REGION Network 37: Validation position reached with module correction
   RUNG wire#powerrail
      Contact( #TMP_xAlwaysON )
      wire#w1
      Contact( #STC_tPZD_Pos.tR.tZSW1.x10 )
      wire#w2
      P_Trig( #STC_tOS_PN.x7 )
      Contact( #STC_tEXT_DATA.tW.xModuleCorrect )
      Contact( #IN_xPositioning )
      { S7_Templates := "SrcType := DInt" } LT_Contact(in1 := #STC_tPROP.d4, in2 := DINT#0)
      S_Coil( #STC_tST.x7 )
   END_RUNG
   RUNG wire#w2
      Contact( #STC_tST.x11 )
      Contact( #STC_tEXT_DATA.tW.xModuleCorrect )
      Contact( #IN_xPositioning )
      { S7_Templates := "SrcType := DInt" } EQ_Contact(in1 := #STC_tPROP.d4, in2 := DINT#0)
      S_Coil( #STC_tST.x7 )
   END_RUNG
   RUNG wire#w1
      I_Contact( #STC_tUSER_DATA.tR.xReadyToMove )
      wire#w3
      R_Coil( #STC_tST.x7 )
   END_RUNG
   RUNG wire#w1
      I_Contact( #IN_xPositioning )
   END_RUNG wire#w3
   RUNG wire#w1
      I_Contact( #STC_tEXT_DATA.tW.xModuleCorrect )
   END_RUNG wire#w3
   RUNG wire#w1
      { S7_Templates := "SrcType := DInt" } GT_Contact(in1 := #STC_tPROP.d4, in2 := DINT#0)
   END_RUNG wire#w3
   // the same network as SCL:
   #_w1 := #TMP_xAlwaysON AND #STC_tPZD_Pos.tR.tZSW1.x10;
   #_w2 := #_w1 AND NOT #STC_tOS_PN.x7;   // rising edge
   #STC_tOS_PN.x7 := #_w1;
   IF #_w2 AND #STC_tEXT_DATA.tW.xModuleCorrect AND #IN_xPositioning AND (#STC_tPROP.d4 < DINT#0) THEN
       #STC_tST.x7 := TRUE;
   END_IF;
   IF #_w1 AND #STC_tST.x11 AND #STC_tEXT_DATA.tW.xModuleCorrect AND #IN_xPositioning AND (#STC_tPROP.d4 = DINT#0) THEN
       #STC_tST.x7 := TRUE;
   END_IF;
   IF #TMP_xAlwaysON AND (NOT #STC_tUSER_DATA.tR.xReadyToMove OR NOT #IN_xPositioning OR NOT #STC_tEXT_DATA.tW.xModuleCorrect OR (#STC_tPROP.d4 > DINT#0)) THEN
       #STC_tST.x7 := FALSE;
   END_IF;
END_REGION

REGION Network 38: Positioning reached
   RUNG wire#powerrail
      Contact( #STC_tUSER_DATA.tR.xReadyToMove )
      Contact( #IN_xPositioning )
      Contact( #STC_tPZD_Pos.tR.tZSW1.x10 )
      wire#w1
      { S7_Templates := "SrcType := DInt" } GE_Contact(in1 := #STC_tPROP.d4, in2 := #TMP_dActualPosMin_cmm)
      { S7_Templates := "SrcType := DInt" } LE_Contact(in1 := #STC_tPROP.d4, in2 := #TMP_dActualPosMax_cmm)
      wire#w2
      Contact( #STC_tPZD_Pos.tR.tPOS_ZSW2.x2 )
      I_Contact( #STC_tPZD_Pos.tR.tPOS_ZSW2.x15 )
      I_Contact( #STC_tPZD_Pos.tW.tSTW1.x6 )
      I_Contact( #STC_tPZD_Pos.tR.tZSW1.x12 )
      Coil( #TMP_x )
   END_RUNG
   RUNG wire#w1
      Contact( #STC_tUSER_DATA.tW.xRelativePosition )
   END_RUNG wire#w2
   RUNG wire#w1
      { S7_Templates := "SrcType := DInt" } LT_Contact(in1 := #STC_tPROP.d4, in2 := 0)
   END_RUNG wire#w2
   RUNG wire#w1
      Contact( #STC_tST.x7 )
   END_RUNG wire#w2
   // the same network as SCL:
   #TMP_x := #STC_tUSER_DATA.tR.xReadyToMove AND #IN_xPositioning AND #STC_tPZD_Pos.tR.tZSW1.x10 AND (((#STC_tPROP.d4 >= #TMP_dActualPosMin_cmm) AND (#STC_tPROP.d4 <= #TMP_dActualPosMax_cmm)) OR #STC_tUSER_DATA.tW.xRelativePosition OR (#STC_tPROP.d4 < 0) OR #STC_tST.x7) AND #STC_tPZD_Pos.tR.tPOS_ZSW2.x2 AND NOT #STC_tPZD_Pos.tR.tPOS_ZSW2.x15 AND NOT #STC_tPZD_Pos.tW.tSTW1.x6 AND NOT #STC_tPZD_Pos.tR.tZSW1.x12;
END_REGION

REGION Network 39: Positioning reached
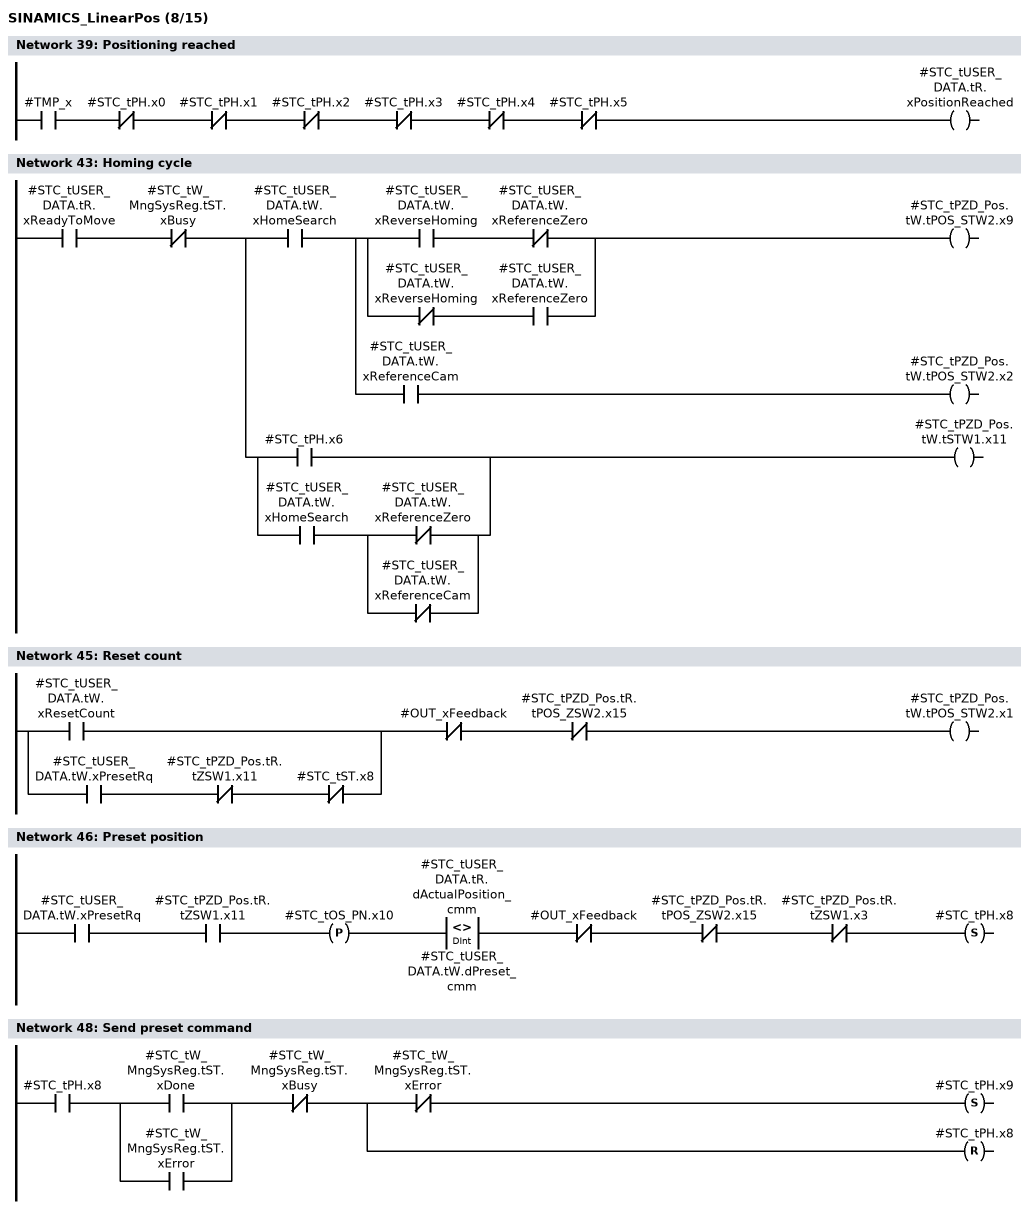
   RUNG wire#powerrail
      Contact( #TMP_x )
      I_Contact( #STC_tPH.x0 )
      I_Contact( #STC_tPH.x1 )
      I_Contact( #STC_tPH.x2 )
      I_Contact( #STC_tPH.x3 )
      I_Contact( #STC_tPH.x4 )
      I_Contact( #STC_tPH.x5 )
      Coil( #STC_tUSER_DATA.tR.xPositionReached )
   END_RUNG
   // the same network as SCL:
   #STC_tUSER_DATA.tR.xPositionReached := #TMP_x AND NOT #STC_tPH.x0 AND NOT #STC_tPH.x1 AND NOT #STC_tPH.x2 AND NOT #STC_tPH.x3 AND NOT #STC_tPH.x4 AND NOT #STC_tPH.x5;
END_REGION

REGION Network 40: #####_HOMING_CYCLE_#####
END_REGION

REGION Network 41 (STL): Send homing preset
         A     #STC_tUSER_DATA.tW.xHomeSearch;
         AN    #STC_tPZD_Pos.tW.tSTW1.x11;
         JCN   PrH0;
         =     #STC_tW_MngSysReg.tST.xWrite_Request;

         L     #STC_tSYS_DATA.iPosPZD_MM;
         SLW   8;
         L     W#16#2;
         OW;
         T     #STC_tW_MngSysReg.tDATA.wRequest_refere_RequestID;
         L     #STC_tSYS_DATA.iPosPZD_MM;
         SLW   8;
         L     W#16#1;
         OW;
         T     #STC_tW_MngSysReg.tDATA.wAxis_NoOfParameters;
         L     W#16#1001;
         T     #STC_tW_MngSysReg.tDATA.wAttribute_NoOfElements;
         L     2599;
         T     #STC_tW_MngSysReg.tDATA.iParameter_number;
         L     W#16#0;
         T     #STC_tW_MngSysReg.tDATA.wSubindex;
         L     W#16#4301;
         T     #STC_tW_MngSysReg.tDATA.wFormat_NoOfValue;
         L     #STC_tSYS_DATA.iDiagAddress;
         T     #STC_tW_MngSysReg.tST.ID;
         L     47;
         T     #STC_tW_MngSysReg.tST.dINDEX;
         L     16;
         T     #STC_tW_MngSysReg.tST.uiLEN;

         L     #STC_tUSER_DATA.tW.dPreset_cmm;
   //      L     DINT#10
   //      *D
         T     #STC_tW_MngSysReg.tDATA.dwRegisterValue;

         CALL  #STC_tWriteRecord
         ( REQ    := #STC_tW_MngSysReg.tST.xWrite_Request,
           ID     := #STC_tW_MngSysReg.tST.ID,
           INDEX  := #STC_tW_MngSysReg.tST.dINDEX,
           LEN    := #STC_tW_MngSysReg.tST.uiLEN,
           DONE   := #STC_tW_MngSysReg.tST.xDone,
           BUSY   := #STC_tW_MngSysReg.tST.xBusy,
           ERROR  := #STC_tW_MngSysReg.tST.xError,
           STATUS := #STC_tW_MngSysReg.tST.dwSTATUS,
           RECORD := #STC_tW_MngSysReg.tDATA
         );
   PrH0: NOP   0;
END_REGION

REGION Network 42 (STL): Error during Send homing preset
         A     #STC_tW_MngSysReg.tST.xError;
         L     34;
         JC    Err;
END_REGION

REGION Network 43: Homing cycle
   RUNG wire#powerrail
      Contact( #STC_tUSER_DATA.tR.xReadyToMove )
      I_Contact( #STC_tW_MngSysReg.tST.xBusy )
      wire#w1
      Contact( #STC_tUSER_DATA.tW.xHomeSearch )
      wire#w2
      Contact( #STC_tUSER_DATA.tW.xReverseHoming )
      I_Contact( #STC_tUSER_DATA.tW.xReferenceZero )
      wire#w3
      Coil( #STC_tPZD_Pos.tW.tPOS_STW2.x9 )
   END_RUNG
   RUNG wire#w2
      I_Contact( #STC_tUSER_DATA.tW.xReverseHoming )
      Contact( #STC_tUSER_DATA.tW.xReferenceZero )
   END_RUNG wire#w3
   RUNG wire#w2
      Contact( #STC_tUSER_DATA.tW.xReferenceCam )
      Coil( #STC_tPZD_Pos.tW.tPOS_STW2.x2 )
   END_RUNG
   RUNG wire#w1
      Contact( #STC_tPH.x6 )
      wire#w4
      Coil( #STC_tPZD_Pos.tW.tSTW1.x11 )
   END_RUNG
   RUNG wire#w1
      Contact( #STC_tUSER_DATA.tW.xHomeSearch )
      wire#w5
      I_Contact( #STC_tUSER_DATA.tW.xReferenceZero )
   END_RUNG wire#w4
   RUNG wire#w5
      I_Contact( #STC_tUSER_DATA.tW.xReferenceCam )
   END_RUNG wire#w4
   // the same network as SCL:
   #_w1 := #STC_tUSER_DATA.tR.xReadyToMove AND NOT #STC_tW_MngSysReg.tST.xBusy;
   #_w2 := #_w1 AND #STC_tUSER_DATA.tW.xHomeSearch;
   #STC_tPZD_Pos.tW.tPOS_STW2.x9 := #_w2 AND ((#STC_tUSER_DATA.tW.xReverseHoming AND NOT #STC_tUSER_DATA.tW.xReferenceZero) OR (NOT #STC_tUSER_DATA.tW.xReverseHoming AND #STC_tUSER_DATA.tW.xReferenceZero));
   #STC_tPZD_Pos.tW.tPOS_STW2.x2 := #_w2 AND #STC_tUSER_DATA.tW.xReferenceCam;
   #STC_tPZD_Pos.tW.tSTW1.x11 := #_w1 AND (#STC_tPH.x6 OR (#STC_tUSER_DATA.tW.xHomeSearch AND (NOT #STC_tUSER_DATA.tW.xReferenceZero OR NOT #STC_tUSER_DATA.tW.xReferenceCam)));
END_REGION

REGION Network 44: #####_PRESET_ACTUAL_POSITION_#####
END_REGION

REGION Network 45: Reset count
   RUNG wire#powerrail
      Contact( #STC_tUSER_DATA.tW.xResetCount )
      wire#w1
      I_Contact( #OUT_xFeedback )
      I_Contact( #STC_tPZD_Pos.tR.tPOS_ZSW2.x15 )
      Coil( #STC_tPZD_Pos.tW.tPOS_STW2.x1 )
   END_RUNG
   RUNG wire#powerrail
      Contact( #STC_tUSER_DATA.tW.xPresetRq )
      I_Contact( #STC_tPZD_Pos.tR.tZSW1.x11 )
      I_Contact( #STC_tST.x8 )
   END_RUNG wire#w1
   // the same network as SCL:
   #STC_tPZD_Pos.tW.tPOS_STW2.x1 := (#STC_tUSER_DATA.tW.xResetCount OR (#STC_tUSER_DATA.tW.xPresetRq AND NOT #STC_tPZD_Pos.tR.tZSW1.x11 AND NOT #STC_tST.x8)) AND NOT #OUT_xFeedback AND NOT #STC_tPZD_Pos.tR.tPOS_ZSW2.x15;
END_REGION

REGION Network 46: Preset position
   RUNG wire#powerrail
      Contact( #STC_tUSER_DATA.tW.xPresetRq )
      Contact( #STC_tPZD_Pos.tR.tZSW1.x11 )
      P_Trig( #STC_tOS_PN.x10 )
      { S7_Templates := "SrcType := DInt" } NE_Contact(in1 := #STC_tUSER_DATA.tR.dActualPosition_cmm, in2 := #STC_tUSER_DATA.tW.dPreset_cmm)
      I_Contact( #OUT_xFeedback )
      I_Contact( #STC_tPZD_Pos.tR.tPOS_ZSW2.x15 )
      I_Contact( #STC_tPZD_Pos.tR.tZSW1.x3 )
      S_Coil( #STC_tPH.x8 )
   END_RUNG
   // the same network as SCL:
   #_w1 := #STC_tUSER_DATA.tW.xPresetRq AND #STC_tPZD_Pos.tR.tZSW1.x11;
   #_w2 := #_w1 AND NOT #STC_tOS_PN.x10;   // rising edge
   #STC_tOS_PN.x10 := #_w1;
   IF #_w2 AND (#STC_tUSER_DATA.tR.dActualPosition_cmm <> #STC_tUSER_DATA.tW.dPreset_cmm) AND NOT #OUT_xFeedback AND NOT #STC_tPZD_Pos.tR.tPOS_ZSW2.x15 AND NOT #STC_tPZD_Pos.tR.tZSW1.x3 THEN
       #STC_tPH.x8 := TRUE;
   END_IF;
END_REGION

REGION Network 47 (STL): Send encoder value
         A     #STC_tPH.x8;
         JCN   PrE0;
         =     #STC_tW_MngSysReg.tST.xWrite_Request;

         L     #STC_tSYS_DATA.iPosPZD_MM;
         +     10;
         SLW   8;
         L     W#16#2;
         OW;
         T     #STC_tW_MngSysReg.tDATA.wRequest_refere_RequestID;
         L     #STC_tSYS_DATA.iPosPZD_MM;
         SLW   8;
         L     W#16#1;
         OW;
         T     #STC_tW_MngSysReg.tDATA.wAxis_NoOfParameters;
         L     W#16#1001;
         T     #STC_tW_MngSysReg.tDATA.wAttribute_NoOfElements;
         L     2599;
         T     #STC_tW_MngSysReg.tDATA.iParameter_number;
         L     W#16#0;
         T     #STC_tW_MngSysReg.tDATA.wSubindex;
         L     W#16#4301;
         T     #STC_tW_MngSysReg.tDATA.wFormat_NoOfValue;
         L     #STC_tSYS_DATA.iDiagAddress;
         T     #STC_tW_MngSysReg.tST.ID;
         L     47;
         T     #STC_tW_MngSysReg.tST.dINDEX;
         L     16;
         T     #STC_tW_MngSysReg.tST.uiLEN;

         L     #STC_tUSER_DATA.tW.dPreset_cmm;
   //  L     DINT#10
   //  *D
         T     #STC_tW_MngSysReg.tDATA.dwRegisterValue;

         CALL  #STC_tWriteRecord
         ( REQ    := #STC_tW_MngSysReg.tST.xWrite_Request,
           ID     := #STC_tW_MngSysReg.tST.ID,
           INDEX  := #STC_tW_MngSysReg.tST.dINDEX,
           LEN    := #STC_tW_MngSysReg.tST.uiLEN,
           DONE   := #STC_tW_MngSysReg.tST.xDone,
           BUSY   := #STC_tW_MngSysReg.tST.xBusy,
           ERROR  := #STC_tW_MngSysReg.tST.xError,
           STATUS := #STC_tW_MngSysReg.tST.dwSTATUS,
           RECORD := #STC_tW_MngSysReg.tDATA
         );
   PrE0: NOP   0;
END_REGION

REGION Network 48: Send preset command
   RUNG wire#powerrail
      Contact( #STC_tPH.x8 )
      wire#w1
      Contact( #STC_tW_MngSysReg.tST.xDone )
      wire#w2
      I_Contact( #STC_tW_MngSysReg.tST.xBusy )
      wire#w3
      I_Contact( #STC_tW_MngSysReg.tST.xError )
      S_Coil( #STC_tPH.x9 )
   END_RUNG
   RUNG wire#w1
      Contact( #STC_tW_MngSysReg.tST.xError )
   END_RUNG wire#w2
   RUNG wire#w3
      R_Coil( #STC_tPH.x8 )
   END_RUNG
   // the same network as SCL:
   #_w1 := #STC_tPH.x8 AND (#STC_tW_MngSysReg.tST.xDone OR #STC_tW_MngSysReg.tST.xError) AND NOT #STC_tW_MngSysReg.tST.xBusy;
   IF #_w1 AND NOT #STC_tW_MngSysReg.tST.xError THEN #STC_tPH.x9 := TRUE; END_IF;
   IF #_w1 THEN #STC_tPH.x8 := FALSE; END_IF;
END_REGION

REGION Network 49 (STL): Error during send ecoder value
         A     #STC_tW_MngSysReg.tST.xError;
         L     30;
         JC    Err;
END_REGION

REGION Network 50 (STL): Send preset command
         A     #STC_tPH.x9;
         JCN   PrE1;
         =     #STC_tW_MngSysReg.tST.xWrite_Request;

         L     #STC_tSYS_DATA.iPosPZD_MM;
         +     20;
         SLW   8;
         L     W#16#2;
         OW;
         T     #STC_tW_MngSysReg.tDATA.wRequest_refere_RequestID;
         L     #STC_tSYS_DATA.iPosPZD_MM;
         SLW   8;
         L     W#16#1;
         OW;
         T     #STC_tW_MngSysReg.tDATA.wAxis_NoOfParameters;
         L     W#16#1001;
         T     #STC_tW_MngSysReg.tDATA.wAttribute_NoOfElements;
         L     2507;
         T     #STC_tW_MngSysReg.tDATA.iParameter_number;
         L     #STC_tSYS_DATA.iEncNumb;
         T     #STC_tW_MngSysReg.tDATA.wSubindex;
         L     W#16#4201;
         T     #STC_tW_MngSysReg.tDATA.wFormat_NoOfValue;
         L     #STC_tSYS_DATA.iDiagAddress;
         T     #STC_tW_MngSysReg.tST.ID;
         L     47;
         T     #STC_tW_MngSysReg.tST.dINDEX;
         L     14;
         T     #STC_tW_MngSysReg.tST.uiLEN;

         L     DINT#2;
         SLD   16;
         T     #STC_tW_MngSysReg.tDATA.dwRegisterValue;

         CALL  #STC_tWriteRecord
         ( REQ    := #STC_tW_MngSysReg.tST.xWrite_Request,
           ID     := #STC_tW_MngSysReg.tST.ID,
           INDEX  := #STC_tW_MngSysReg.tST.dINDEX,
           LEN    := #STC_tW_MngSysReg.tST.uiLEN,
           DONE   := #STC_tW_MngSysReg.tST.xDone,
           BUSY   := #STC_tW_MngSysReg.tST.xBusy,
           ERROR  := #STC_tW_MngSysReg.tST.xError,
           STATUS := #STC_tW_MngSysReg.tST.dwSTATUS,
           RECORD := #STC_tW_MngSysReg.tDATA
         );
   PrE1: NOP   0;
END_REGION

REGION Network 51: Send saving preset command
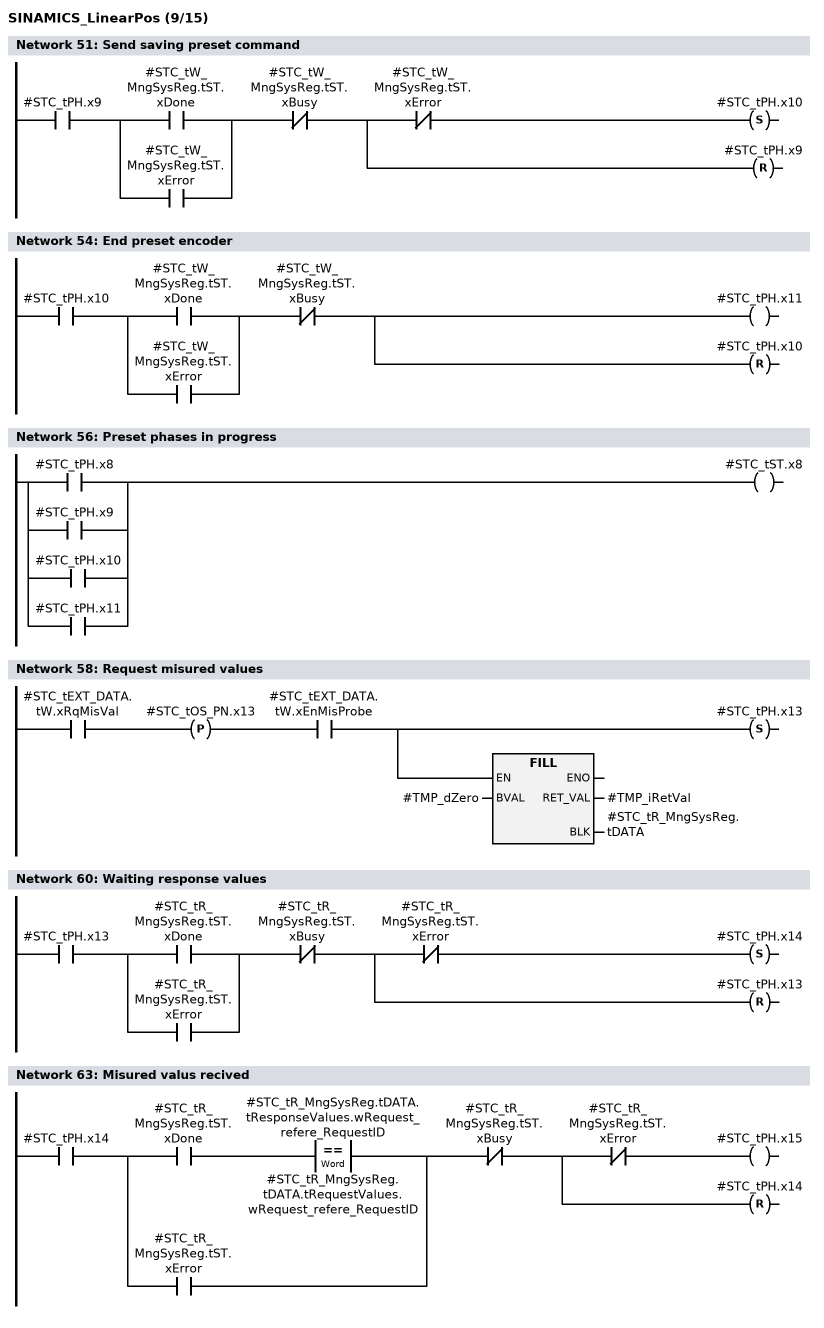
   RUNG wire#powerrail
      Contact( #STC_tPH.x9 )
      wire#w1
      Contact( #STC_tW_MngSysReg.tST.xDone )
      wire#w2
      I_Contact( #STC_tW_MngSysReg.tST.xBusy )
      wire#w3
      I_Contact( #STC_tW_MngSysReg.tST.xError )
      S_Coil( #STC_tPH.x10 )
   END_RUNG
   RUNG wire#w1
      Contact( #STC_tW_MngSysReg.tST.xError )
   END_RUNG wire#w2
   RUNG wire#w3
      R_Coil( #STC_tPH.x9 )
   END_RUNG
   // the same network as SCL:
   #_w1 := #STC_tPH.x9 AND (#STC_tW_MngSysReg.tST.xDone OR #STC_tW_MngSysReg.tST.xError) AND NOT #STC_tW_MngSysReg.tST.xBusy;
   IF #_w1 AND NOT #STC_tW_MngSysReg.tST.xError THEN #STC_tPH.x10 := TRUE; END_IF;
   IF #_w1 THEN #STC_tPH.x9 := FALSE; END_IF;
END_REGION

REGION Network 52 (STL): Error during preset command
         A     #STC_tW_MngSysReg.tST.xError;
         L     31;
         JC    Err;
END_REGION

REGION Network 53 (STL): Send saving preset command
         A     #STC_tPH.x10;
         JCN   PrE2;
         =     #STC_tW_MngSysReg.tST.xWrite_Request;

         L     #STC_tSYS_DATA.iPosPZD_MM;
         +     30;
         SLW   8;
         L     W#16#2;
         OW;
         T     #STC_tW_MngSysReg.tDATA.wRequest_refere_RequestID;
         L     #STC_tSYS_DATA.iPosPZD_CU;
         SLW   8;
         L     W#16#1;
         OW;
         T     #STC_tW_MngSysReg.tDATA.wAxis_NoOfParameters;
         L     W#16#1001;
         T     #STC_tW_MngSysReg.tDATA.wAttribute_NoOfElements;
         L     977;
         T     #STC_tW_MngSysReg.tDATA.iParameter_number;
         L     W#16#0;
         T     #STC_tW_MngSysReg.tDATA.wSubindex;
         L     W#16#4201;
         T     #STC_tW_MngSysReg.tDATA.wFormat_NoOfValue;
         L     #STC_tSYS_DATA.iDiagAddress;
         T     #STC_tW_MngSysReg.tST.ID;
         L     47;
         T     #STC_tW_MngSysReg.tST.dINDEX;
         L     14;
         T     #STC_tW_MngSysReg.tST.uiLEN;

         L     DINT#1;
         SLD   16;
         T     #STC_tW_MngSysReg.tDATA.dwRegisterValue;

         CALL  #STC_tWriteRecord
         ( REQ    := #STC_tW_MngSysReg.tST.xWrite_Request,
           ID     := #STC_tW_MngSysReg.tST.ID,
           INDEX  := #STC_tW_MngSysReg.tST.dINDEX,
           LEN    := #STC_tW_MngSysReg.tST.uiLEN,
           DONE   := #STC_tW_MngSysReg.tST.xDone,
           BUSY   := #STC_tW_MngSysReg.tST.xBusy,
           ERROR  := #STC_tW_MngSysReg.tST.xError,
           STATUS := #STC_tW_MngSysReg.tST.dwSTATUS,
           RECORD := #STC_tW_MngSysReg.tDATA
         );
   PrE2: NOP   0;
END_REGION

REGION Network 54: End preset encoder
   RUNG wire#powerrail
      Contact( #STC_tPH.x10 )
      wire#w1
      Contact( #STC_tW_MngSysReg.tST.xDone )
      wire#w2
      I_Contact( #STC_tW_MngSysReg.tST.xBusy )
      wire#w3
      Coil( #STC_tPH.x11 )
   END_RUNG
   RUNG wire#w1
      Contact( #STC_tW_MngSysReg.tST.xError )
   END_RUNG wire#w2
   RUNG wire#w3
      R_Coil( #STC_tPH.x10 )
   END_RUNG
   // the same network as SCL:
   #STC_tPH.x11 := #STC_tPH.x10 AND (#STC_tW_MngSysReg.tST.xDone OR #STC_tW_MngSysReg.tST.xError) AND NOT #STC_tW_MngSysReg.tST.xBusy;
   IF #STC_tPH.x11 THEN #STC_tPH.x10 := FALSE; END_IF;
END_REGION

REGION Network 55 (STL): Error during saving preset command
         A     #STC_tW_MngSysReg.tST.xError;
         L     32;
         JC    Err;
END_REGION

REGION Network 56: Preset phases in progress
   RUNG wire#powerrail
      Contact( #STC_tPH.x8 )
      wire#w1
      Coil( #STC_tST.x8 )
   END_RUNG
   RUNG wire#powerrail
      Contact( #STC_tPH.x9 )
   END_RUNG wire#w1
   RUNG wire#powerrail
      Contact( #STC_tPH.x10 )
   END_RUNG wire#w1
   RUNG wire#powerrail
      Contact( #STC_tPH.x11 )
   END_RUNG wire#w1
   // the same network as SCL:
   #STC_tST.x8 := #STC_tPH.x8 OR #STC_tPH.x9 OR #STC_tPH.x10 OR #STC_tPH.x11;
END_REGION

REGION Network 57: #####_READING_MISURED_VALUES_#####
END_REGION

REGION Network 58: Request misured values
   #_w1 := #STC_tEXT_DATA.tW.xRqMisVal AND NOT #STC_tOS_PN.x13;   // rising edge
   #STC_tOS_PN.x13 := #STC_tEXT_DATA.tW.xRqMisVal;
   IF #_w1 AND #STC_tEXT_DATA.tW.xEnMisProbe THEN
       #STC_tPH.x13 := TRUE;
       #TMP_iRetVal := FILL(BVAL := #TMP_dZero, BLK => #STC_tR_MngSysReg.tDATA);
   END_IF;
END_REGION

REGION Network 59 (STL): Send request misured values
         A     #STC_tPH.x13;
         JCN   RdV1;
         =     #STC_tR_MngSysReg.tST.xRead_Request;

         L     #STC_tSYS_DATA.iPosPZD_MM;
         +     40;
         SLW   8;
         L     W#16#1;
         OW;
         T     #STC_tR_MngSysReg.tDATA.tRequestValues.wRequest_refere_RequestID;
         L     #STC_tSYS_DATA.iPosPZD_MM;
         SLW   8;
         L     W#16#C;
         OW;
         T     #STC_tR_MngSysReg.tDATA.tRequestValues.wAxis_NoOfParameters;
         L     W#16#1000;
         T     #STC_tR_MngSysReg.tDATA.tRequestValues.wAttribute_NoOfElements_1;
         L     21700;
         T     #STC_tR_MngSysReg.tDATA.tRequestValues.iParameter_number_1;
         L     W#16#0;
         T     #STC_tR_MngSysReg.tDATA.tRequestValues.wSubindex_1;

         L     W#16#1000;
         T     #STC_tR_MngSysReg.tDATA.tRequestValues.wAttribute_NoOfElements_2;
         L     21701;
         T     #STC_tR_MngSysReg.tDATA.tRequestValues.iParameter_number_2;
         L     W#16#0;
         T     #STC_tR_MngSysReg.tDATA.tRequestValues.wSubindex_2;

         L     W#16#1000;
         T     #STC_tR_MngSysReg.tDATA.tRequestValues.wAttribute_NoOfElements_3;
         L     21702;
         T     #STC_tR_MngSysReg.tDATA.tRequestValues.iParameter_number_3;
         L     W#16#0;
         T     #STC_tR_MngSysReg.tDATA.tRequestValues.wSubindex_3;

         L     W#16#1000;
         T     #STC_tR_MngSysReg.tDATA.tRequestValues.wAttribute_NoOfElements_4;
         L     21703;
         T     #STC_tR_MngSysReg.tDATA.tRequestValues.iParameter_number_4;
         L     W#16#0;
         T     #STC_tR_MngSysReg.tDATA.tRequestValues.wSubindex_4;

         L     W#16#1000;
         T     #STC_tR_MngSysReg.tDATA.tRequestValues.wAttribute_NoOfElements_5;
         L     21704;
         T     #STC_tR_MngSysReg.tDATA.tRequestValues.iParameter_number_5;
         L     W#16#0;
         T     #STC_tR_MngSysReg.tDATA.tRequestValues.wSubindex_5;

         L     W#16#1000;
         T     #STC_tR_MngSysReg.tDATA.tRequestValues.wAttribute_NoOfElements_6;
         L     21705;
         T     #STC_tR_MngSysReg.tDATA.tRequestValues.iParameter_number_6;
         L     W#16#0;
         T     #STC_tR_MngSysReg.tDATA.tRequestValues.wSubindex_6;

         L     W#16#1000;
         T     #STC_tR_MngSysReg.tDATA.tRequestValues.wAttribute_NoOfElements_7;
         L     21712;
         T     #STC_tR_MngSysReg.tDATA.tRequestValues.iParameter_number_7;
         L     W#16#0;
         T     #STC_tR_MngSysReg.tDATA.tRequestValues.wSubindex_7;

         L     W#16#1000;
         T     #STC_tR_MngSysReg.tDATA.tRequestValues.wAttribute_NoOfElements_8;
         L     21713;
         T     #STC_tR_MngSysReg.tDATA.tRequestValues.iParameter_number_8;
         L     W#16#0;
         T     #STC_tR_MngSysReg.tDATA.tRequestValues.wSubindex_8;

         L     W#16#1000;
         T     #STC_tR_MngSysReg.tDATA.tRequestValues.wAttribute_NoOfElements_9;
         L     21714;
         T     #STC_tR_MngSysReg.tDATA.tRequestValues.iParameter_number_9;
         L     W#16#0;
         T     #STC_tR_MngSysReg.tDATA.tRequestValues.wSubindex_9;

         L     W#16#1000;
         T     #STC_tR_MngSysReg.tDATA.tRequestValues.wAttribute_NoOfElement_10;
         L     21715;
         T     #STC_tR_MngSysReg.tDATA.tRequestValues.iParameter_number_10;
         L     W#16#0;
         T     #STC_tR_MngSysReg.tDATA.tRequestValues.wSubindex_10;

         L     W#16#1000;
         T     #STC_tR_MngSysReg.tDATA.tRequestValues.wAttribute_NoOfElement_11;
         L     21716;
         T     #STC_tR_MngSysReg.tDATA.tRequestValues.iParameter_number_11;
         L     W#16#0;
         T     #STC_tR_MngSysReg.tDATA.tRequestValues.wSubindex_11;

         L     W#16#1000;
         T     #STC_tR_MngSysReg.tDATA.tRequestValues.wAttribute_NoOfElement_12;
         L     21717;
         T     #STC_tR_MngSysReg.tDATA.tRequestValues.iParameter_number_12;
         L     W#16#0;
         T     #STC_tR_MngSysReg.tDATA.tRequestValues.wSubindex_12;

         L     #STC_tSYS_DATA.iDiagAddress;
         T     #STC_tR_MngSysReg.tST.ID;
         L     47;
         T     #STC_tR_MngSysReg.tST.dINDEX;
         L     76;
         T     #STC_tR_MngSysReg.tST.uiLEN;

         CALL  #STC_tWriteRecord
         ( REQ    := #STC_tR_MngSysReg.tST.xRead_Request,
           ID     := #STC_tR_MngSysReg.tST.ID,
           INDEX  := #STC_tR_MngSysReg.tST.dINDEX,
           LEN    := #STC_tR_MngSysReg.tST.uiLEN,
           DONE   := #STC_tR_MngSysReg.tST.xDone,
           BUSY   := #STC_tR_MngSysReg.tST.xBusy,
           ERROR  := #STC_tR_MngSysReg.tST.xError,
           STATUS := #STC_tR_MngSysReg.tST.dwSTATUS,
           RECORD := #STC_tR_MngSysReg.tDATA.tRequestValues
         );

   RdV1: NOP   0;
END_REGION

REGION Network 60: Waiting response values
   RUNG wire#powerrail
      Contact( #STC_tPH.x13 )
      wire#w1
      Contact( #STC_tR_MngSysReg.tST.xDone )
      wire#w2
      I_Contact( #STC_tR_MngSysReg.tST.xBusy )
      wire#w3
      I_Contact( #STC_tR_MngSysReg.tST.xError )
      S_Coil( #STC_tPH.x14 )
   END_RUNG
   RUNG wire#w1
      Contact( #STC_tR_MngSysReg.tST.xError )
   END_RUNG wire#w2
   RUNG wire#w3
      R_Coil( #STC_tPH.x13 )
   END_RUNG
   // the same network as SCL:
   #_w1 := #STC_tPH.x13 AND (#STC_tR_MngSysReg.tST.xDone OR #STC_tR_MngSysReg.tST.xError) AND NOT #STC_tR_MngSysReg.tST.xBusy;
   IF #_w1 AND NOT #STC_tR_MngSysReg.tST.xError THEN #STC_tPH.x14 := TRUE; END_IF;
   IF #_w1 THEN #STC_tPH.x13 := FALSE; END_IF;
END_REGION

REGION Network 61 (STL): Error during waiting response values
         A     #STC_tR_MngSysReg.tST.xError;
         L     40;
         JC    Err;
END_REGION

REGION Network 62 (STL): Send response misured values
         A     #STC_tPH.x14;
         JCN   RdV2;
         AN    #STC_tR_MngSysReg.tST.xBusy;
         =     #STC_tR_MngSysReg.tST.xRead_Request;

         L     #STC_tSYS_DATA.iDiagAddress;
         T     #STC_tR_MngSysReg.tST.ID;
         L     47;
         T     #STC_tR_MngSysReg.tST.dINDEX;
         L     76;
         T     #STC_tR_MngSysReg.tST.uiMLEN;

         CALL  #STC_tReadRecord
         ( REQ    := #STC_tR_MngSysReg.tST.xRead_Request,
           ID     := #STC_tR_MngSysReg.tST.ID,
           INDEX  := #STC_tR_MngSysReg.tST.dINDEX,
           MLEN   := #STC_tR_MngSysReg.tST.uiMLEN,
           VALID  := #STC_tR_MngSysReg.tST.xDone,
           BUSY   := #STC_tR_MngSysReg.tST.xBusy,
           ERROR  := #STC_tR_MngSysReg.tST.xError,
           STATUS := #STC_tR_MngSysReg.tST.dwSTATUS,
           LEN    := #STC_tR_MngSysReg.tST.uiLEN,
           RECORD := #STC_tR_MngSysReg.tDATA.tResponseValues
         );

         L     #STC_tR_MngSysReg.tDATA.tResponseValues.wRequest_refere_RequestID;
         L     W#16#FF7F;
         AW;
         T     #STC_tR_MngSysReg.tDATA.tResponseValues.wRequest_refere_RequestID;

   RdV2: NOP   0;
END_REGION

REGION Network 63: Misured valus recived
   RUNG wire#powerrail
      Contact( #STC_tPH.x14 )
      wire#w1
      Contact( #STC_tR_MngSysReg.tST.xDone )
      { S7_Templates := "SrcType := Word" } EQ_Contact(in1 := #STC_tR_MngSysReg.tDATA.tResponseValues.wRequest_refere_RequestID, in2 := #STC_tR_MngSysReg.tDATA.tRequestValues.wRequest_refere_RequestID)
      wire#w2
      I_Contact( #STC_tR_MngSysReg.tST.xBusy )
      wire#w3
      I_Contact( #STC_tR_MngSysReg.tST.xError )
      Coil( #STC_tPH.x15 )
   END_RUNG
   RUNG wire#w1
      Contact( #STC_tR_MngSysReg.tST.xError )
   END_RUNG wire#w2
   RUNG wire#w3
      R_Coil( #STC_tPH.x14 )
   END_RUNG
   // the same network as SCL:
   #_w1 := #STC_tPH.x14 AND ((#STC_tR_MngSysReg.tST.xDone AND (#STC_tR_MngSysReg.tDATA.tResponseValues.wRequest_refere_RequestID = #STC_tR_MngSysReg.tDATA.tRequestValues.wRequest_refere_RequestID)) OR #STC_tR_MngSysReg.tST.xError) AND NOT #STC_tR_MngSysReg.tST.xBusy;
   #STC_tPH.x15 := #_w1 AND NOT #STC_tR_MngSysReg.tST.xError;
   IF #_w1 THEN #STC_tPH.x14 := FALSE; END_IF;
END_REGION

REGION Network 64 (STL): Error during misured valus recived
         A     #STC_tR_MngSysReg.tST.xError;
         L     41;
         JC    Err;
END_REGION

REGION Network 65: Save data
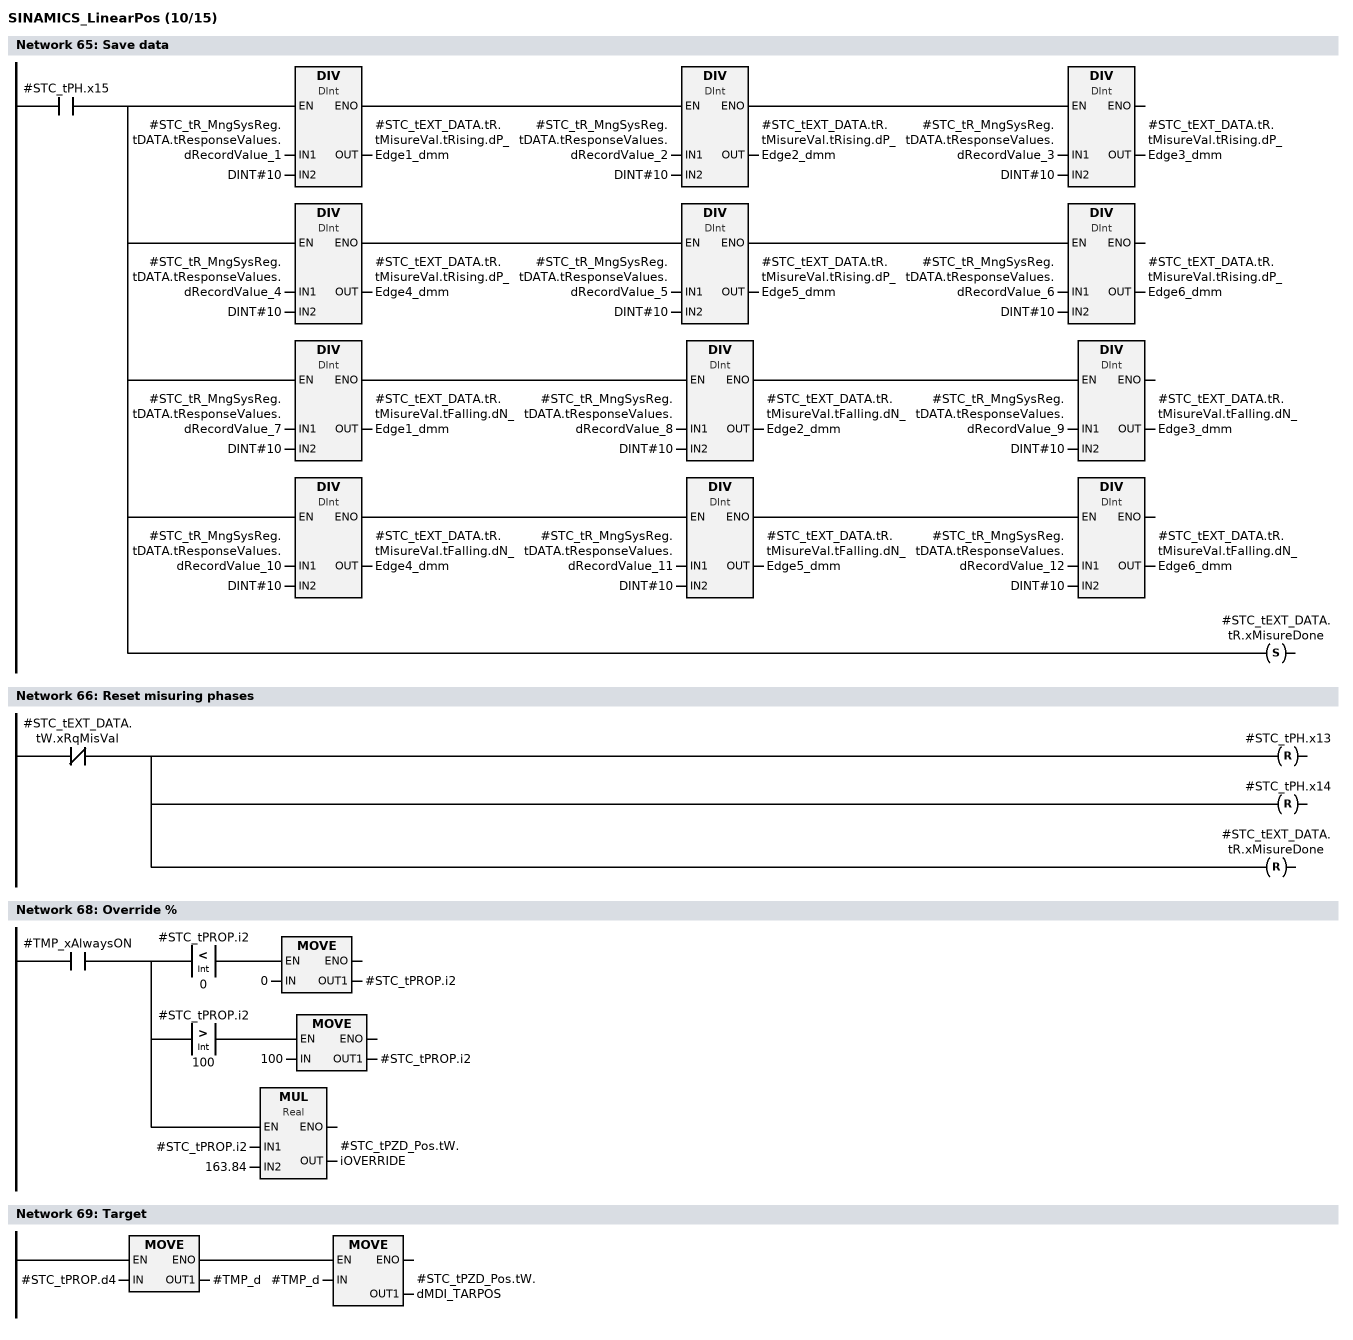
   RUNG wire#powerrail
      Contact( #STC_tPH.x15 )
      wire#w1
      { S7_Templates := "SrcType := DInt"; S7_GenerateENO := "TRUE" } Div(in1 := #STC_tR_MngSysReg.tDATA.tResponseValues.dRecordValue_1, in2 := DINT#10, out => #STC_tEXT_DATA.tR.tMisureVal.tRising.dP_Edge1_dmm)
      { S7_Templates := "SrcType := DInt"; S7_GenerateENO := "TRUE" } Div(in1 := #STC_tR_MngSysReg.tDATA.tResponseValues.dRecordValue_2, in2 := DINT#10, out => #STC_tEXT_DATA.tR.tMisureVal.tRising.dP_Edge2_dmm)
      { S7_Templates := "SrcType := DInt"; S7_GenerateENO := "TRUE" } Div(in1 := #STC_tR_MngSysReg.tDATA.tResponseValues.dRecordValue_3, in2 := DINT#10, out => #STC_tEXT_DATA.tR.tMisureVal.tRising.dP_Edge3_dmm)
   END_RUNG
   RUNG wire#w1
      { S7_Templates := "SrcType := DInt"; S7_GenerateENO := "TRUE" } Div(in1 := #STC_tR_MngSysReg.tDATA.tResponseValues.dRecordValue_4, in2 := DINT#10, out => #STC_tEXT_DATA.tR.tMisureVal.tRising.dP_Edge4_dmm)
      { S7_Templates := "SrcType := DInt"; S7_GenerateENO := "TRUE" } Div(in1 := #STC_tR_MngSysReg.tDATA.tResponseValues.dRecordValue_5, in2 := DINT#10, out => #STC_tEXT_DATA.tR.tMisureVal.tRising.dP_Edge5_dmm)
      { S7_Templates := "SrcType := DInt"; S7_GenerateENO := "TRUE" } Div(in1 := #STC_tR_MngSysReg.tDATA.tResponseValues.dRecordValue_6, in2 := DINT#10, out => #STC_tEXT_DATA.tR.tMisureVal.tRising.dP_Edge6_dmm)
   END_RUNG
   RUNG wire#w1
      { S7_Templates := "SrcType := DInt"; S7_GenerateENO := "TRUE" } Div(in1 := #STC_tR_MngSysReg.tDATA.tResponseValues.dRecordValue_7, in2 := DINT#10, out => #STC_tEXT_DATA.tR.tMisureVal.tFalling.dN_Edge1_dmm)
      { S7_Templates := "SrcType := DInt"; S7_GenerateENO := "TRUE" } Div(in1 := #STC_tR_MngSysReg.tDATA.tResponseValues.dRecordValue_8, in2 := DINT#10, out => #STC_tEXT_DATA.tR.tMisureVal.tFalling.dN_Edge2_dmm)
      { S7_Templates := "SrcType := DInt"; S7_GenerateENO := "TRUE" } Div(in1 := #STC_tR_MngSysReg.tDATA.tResponseValues.dRecordValue_9, in2 := DINT#10, out => #STC_tEXT_DATA.tR.tMisureVal.tFalling.dN_Edge3_dmm)
   END_RUNG
   RUNG wire#w1
      { S7_Templates := "SrcType := DInt"; S7_GenerateENO := "TRUE" } Div(in1 := #STC_tR_MngSysReg.tDATA.tResponseValues.dRecordValue_10, in2 := DINT#10, out => #STC_tEXT_DATA.tR.tMisureVal.tFalling.dN_Edge4_dmm)
      { S7_Templates := "SrcType := DInt"; S7_GenerateENO := "TRUE" } Div(in1 := #STC_tR_MngSysReg.tDATA.tResponseValues.dRecordValue_11, in2 := DINT#10, out => #STC_tEXT_DATA.tR.tMisureVal.tFalling.dN_Edge5_dmm)
      { S7_Templates := "SrcType := DInt"; S7_GenerateENO := "TRUE" } Div(in1 := #STC_tR_MngSysReg.tDATA.tResponseValues.dRecordValue_12, in2 := DINT#10, out => #STC_tEXT_DATA.tR.tMisureVal.tFalling.dN_Edge6_dmm)
   END_RUNG
   RUNG wire#w1
      S_Coil( #STC_tEXT_DATA.tR.xMisureDone )
   END_RUNG
   // the same network as SCL:
   // ENO of a box is taken as its EN; it also drops when the box reports an error
   IF #STC_tPH.x15 THEN
       #STC_tEXT_DATA.tR.tMisureVal.tRising.dP_Edge1_dmm := #STC_tR_MngSysReg.tDATA.tResponseValues.dRecordValue_1 / DINT#10;
       #STC_tEXT_DATA.tR.tMisureVal.tRising.dP_Edge2_dmm := #STC_tR_MngSysReg.tDATA.tResponseValues.dRecordValue_2 / DINT#10;
       #STC_tEXT_DATA.tR.tMisureVal.tRising.dP_Edge3_dmm := #STC_tR_MngSysReg.tDATA.tResponseValues.dRecordValue_3 / DINT#10;
       #STC_tEXT_DATA.tR.tMisureVal.tRising.dP_Edge4_dmm := #STC_tR_MngSysReg.tDATA.tResponseValues.dRecordValue_4 / DINT#10;
       #STC_tEXT_DATA.tR.tMisureVal.tRising.dP_Edge5_dmm := #STC_tR_MngSysReg.tDATA.tResponseValues.dRecordValue_5 / DINT#10;
       #STC_tEXT_DATA.tR.tMisureVal.tRising.dP_Edge6_dmm := #STC_tR_MngSysReg.tDATA.tResponseValues.dRecordValue_6 / DINT#10;
       #STC_tEXT_DATA.tR.tMisureVal.tFalling.dN_Edge1_dmm := #STC_tR_MngSysReg.tDATA.tResponseValues.dRecordValue_7 / DINT#10;
       #STC_tEXT_DATA.tR.tMisureVal.tFalling.dN_Edge2_dmm := #STC_tR_MngSysReg.tDATA.tResponseValues.dRecordValue_8 / DINT#10;
       #STC_tEXT_DATA.tR.tMisureVal.tFalling.dN_Edge3_dmm := #STC_tR_MngSysReg.tDATA.tResponseValues.dRecordValue_9 / DINT#10;
       #STC_tEXT_DATA.tR.tMisureVal.tFalling.dN_Edge4_dmm := #STC_tR_MngSysReg.tDATA.tResponseValues.dRecordValue_10 / DINT#10;
       #STC_tEXT_DATA.tR.tMisureVal.tFalling.dN_Edge5_dmm := #STC_tR_MngSysReg.tDATA.tResponseValues.dRecordValue_11 / DINT#10;
       #STC_tEXT_DATA.tR.tMisureVal.tFalling.dN_Edge6_dmm := #STC_tR_MngSysReg.tDATA.tResponseValues.dRecordValue_12 / DINT#10;
       #STC_tEXT_DATA.tR.xMisureDone := TRUE;
   END_IF;
END_REGION

REGION Network 66: Reset misuring phases
   RUNG wire#powerrail
      I_Contact( #STC_tEXT_DATA.tW.xRqMisVal )
      wire#w1
      R_Coil( #STC_tPH.x13 )
   END_RUNG
   RUNG wire#w1
      R_Coil( #STC_tPH.x14 )
   END_RUNG
   RUNG wire#w1
      R_Coil( #STC_tEXT_DATA.tR.xMisureDone )
   END_RUNG
   // the same network as SCL:
   IF NOT #STC_tEXT_DATA.tW.xRqMisVal THEN
       #STC_tPH.x13 := FALSE;
       #STC_tPH.x14 := FALSE;
       #STC_tEXT_DATA.tR.xMisureDone := FALSE;
   END_IF;
END_REGION

REGION Network 67: #####_PARAMETERS_#####
END_REGION

REGION Network 68: Override %
   RUNG wire#powerrail
      Contact( #TMP_xAlwaysON )
      wire#w1
      { S7_Templates := "SrcType := Int" } LT_Contact(in1 := #STC_tPROP.i2, in2 := 0)
      Move(in := 0, out1 => #STC_tPROP.i2)
   END_RUNG
   RUNG wire#w1
      { S7_Templates := "SrcType := Int" } GT_Contact(in1 := #STC_tPROP.i2, in2 := 100)
      Move(in := 100, out1 => #STC_tPROP.i2)
   END_RUNG
   RUNG wire#w1
      { S7_Templates := "SrcType := Real" } Mul(in1 := #STC_tPROP.i2, in2 := 163.84, out => #STC_tPZD_Pos.tW.iOVERRIDE)
   END_RUNG
   // the same network as SCL:
   IF #TMP_xAlwaysON AND (#STC_tPROP.i2 < 0) THEN #STC_tPROP.i2 := 0; END_IF;
   IF #TMP_xAlwaysON AND (#STC_tPROP.i2 > 100) THEN #STC_tPROP.i2 := 100; END_IF;
   IF #TMP_xAlwaysON THEN #STC_tPZD_Pos.tW.iOVERRIDE := #STC_tPROP.i2 * 163.84; END_IF;
END_REGION

REGION Network 69: Target
   RUNG wire#powerrail
      { S7_GenerateENO := "TRUE" } Move(in := #STC_tPROP.d4, out1 => #TMP_d)
      Move(in := #TMP_d, out1 => #STC_tPZD_Pos.tW.dMDI_TARPOS)
   END_RUNG
   // the same network as SCL:
   // ENO of a box is taken as its EN; it also drops when the box reports an error
   #TMP_d := #STC_tPROP.d4;
   #STC_tPZD_Pos.tW.dMDI_TARPOS := #TMP_d;
END_REGION

REGION Network 70: Speed